REGION Network 6: 2 -Op2- - Reparare palete Zona A
   #f[#_op2](sA := #_nop0,   // "sta"
             nrs := #_op2,
             sB := #_cen,
             iA := "DB2_WORK_BITS".Transport_Conveyor_SQs.SQ_Repaired_Pallet[0] AND #tmr[5].Q,
             cEvac := NOT "x".evac[2],
             iAr := NOT "DB2_WORK_BITS".Transport_Conveyor_SQs.SQ_Repaired_Pallet[0],
             iB := "SCentrorMemT",
             cmdB => #tranzit[#_op2],
             ENO => #_w1);
   #f[2].condRetract := #_w1;
   #f[2].WrkDn := #_w1;
   #f[2].disAlm_apar := #_w1;
   #tmr[5].TON(IN := "DB2_WORK_BITS".Transport_Conveyor_SQs.SQ_Repaired_Pallet[0], PT := T#2s);
END_REGION

REGION Network 7: stoper op
   RUNG wire#powerrail
      Contact( "DB2_WORK_BITS".Transport_Conveyor_SQs.SQ_Repaired_Pallet[0] )
      wire#w1
      Coil( "O".StopReqUp1 )
   END_RUNG
   RUNG wire#powerrail
      Contact( #tranzit[#_op2] )
   END_RUNG wire#w1
   // the same network as SCL:
   "O".StopReqUp1 := "DB2_WORK_BITS".Transport_Conveyor_SQs.SQ_Repaired_Pallet[0] OR #tranzit[#_op2];
END_REGION

REGION Network 8
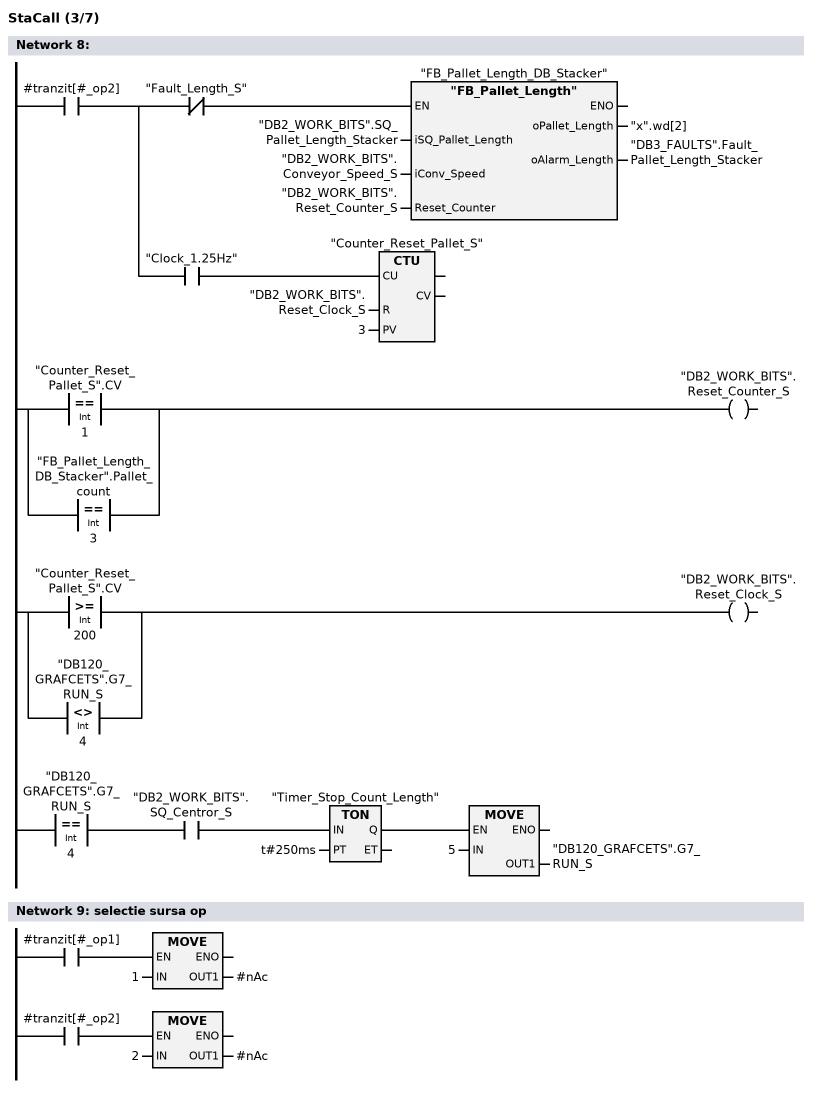
   IF #tranzit[#_op2] AND NOT "Fault_Length_S" THEN
       "FB_Pallet_Length_DB_Stacker"(iSQ_Pallet_Length := "DB2_WORK_BITS".SQ_Pallet_Length_Stacker,   // "FB_Pallet_Length"
                               iConv_Speed := "DB2_WORK_BITS".Conveyor_Speed_S,
                               Reset_Counter := "DB2_WORK_BITS".Reset_Counter_S,
                               oPallet_Length => "x".wd[2],
                               oAlarm_Length => "DB3_FAULTS".Fault_Pallet_Length_Stacker);
   END_IF;
   "Counter_Reset_Pallet_S".CTU(CU := #tranzit[#_op2] AND "Clock_1.25Hz",
                           R := "DB2_WORK_BITS".Reset_Clock_S,
                           PV := 3);
   "DB2_WORK_BITS".Reset_Counter_S := ("Counter_Reset_Pallet_S".CV = 1) OR ("FB_Pallet_Length_DB_Stacker".Pallet_count = 3);
   "DB2_WORK_BITS".Reset_Clock_S := ("Counter_Reset_Pallet_S".CV >= 200) OR ("DB120_GRAFCETS".G7_RUN_S <> 4);
   "Timer_Stop_Count_Length".TON(IN := ("DB120_GRAFCETS".G7_RUN_S = 4) AND "DB2_WORK_BITS".SQ_Centror_S,
                           PT := t#250ms);
   IF "Timer_Stop_Count_Length".Q THEN "DB120_GRAFCETS".G7_RUN_S := 5; END_IF;
END_REGION

REGION Network 9: selectie sursa op
   RUNG wire#powerrail
      Contact( #tranzit[#_op1] )
      Move(in := 1, out1 => #nAc)
   END_RUNG
   RUNG wire#powerrail
      Contact( #tranzit[#_op2] )
      Move(in := 2, out1 => #nAc)
   END_RUNG
   // the same network as SCL:
   IF #tranzit[#_op1] THEN #nAc := 1; END_IF;
   IF #tranzit[#_op2] THEN #nAc := 2; END_IF;
END_REGION

REGION Network 10: senz stop stk
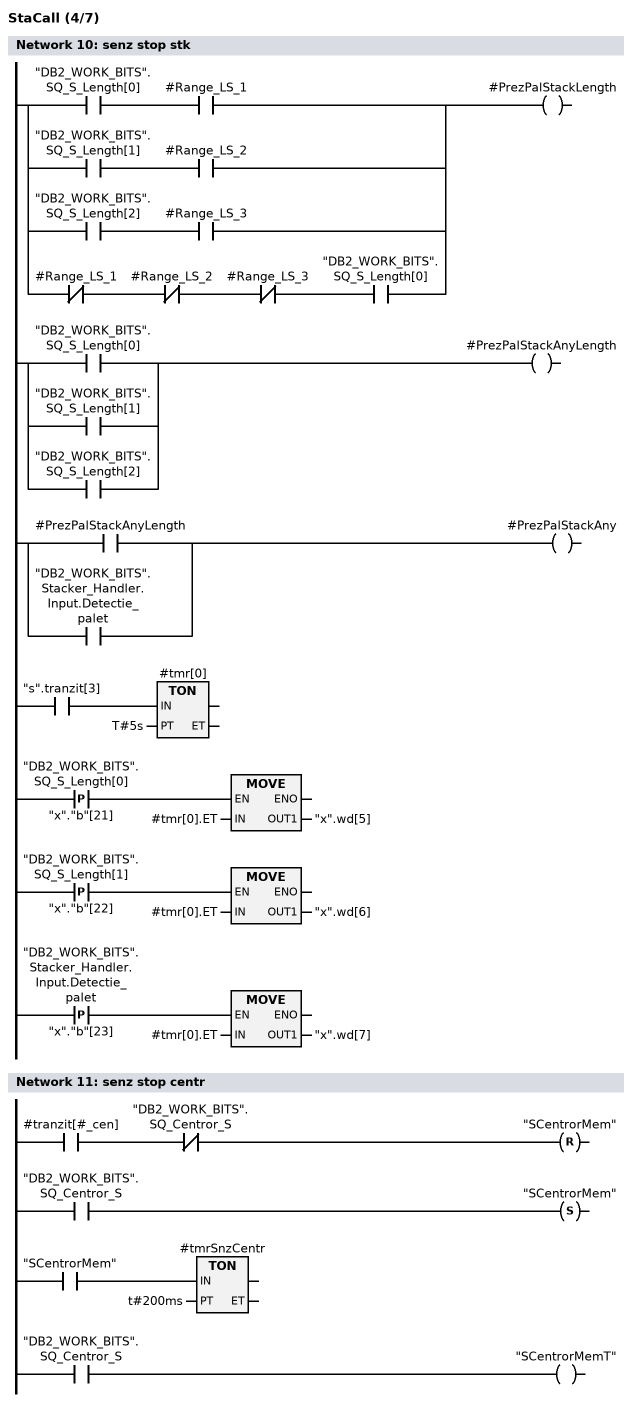
   #PrezPalStackLength := ("DB2_WORK_BITS".SQ_S_Length[0] AND #Range_LS_1) OR ("DB2_WORK_BITS".SQ_S_Length[1] AND #Range_LS_2) OR ("DB2_WORK_BITS".SQ_S_Length[2] AND #Range_LS_3) OR (NOT #Range_LS_1 AND NOT #Range_LS_2 AND NOT #Range_LS_3 AND "DB2_WORK_BITS".SQ_S_Length[0]);
   #PrezPalStackAnyLength := "DB2_WORK_BITS".SQ_S_Length[0] OR "DB2_WORK_BITS".SQ_S_Length[1] OR "DB2_WORK_BITS".SQ_S_Length[2];
   #PrezPalStackAny := #PrezPalStackAnyLength OR "DB2_WORK_BITS".Stacker_Handler.Input.Detectie_palet;
   #tmr[0].TON(IN := "s".tranzit[3], PT := T#5s);
   #_w1 := "DB2_WORK_BITS".SQ_S_Length[0] AND NOT "x"."b"[21];   // rising edge of "DB2_WORK_BITS".SQ_S_Length[0]
   "x"."b"[21] := "DB2_WORK_BITS".SQ_S_Length[0];
   IF #_w1 THEN "x".wd[5] := #tmr[0].ET; END_IF;
   #_w2 := "DB2_WORK_BITS".SQ_S_Length[1] AND NOT "x"."b"[22];   // rising edge of "DB2_WORK_BITS".SQ_S_Length[1]
   "x"."b"[22] := "DB2_WORK_BITS".SQ_S_Length[1];
   IF #_w2 THEN "x".wd[6] := #tmr[0].ET; END_IF;
   #_w3 := "DB2_WORK_BITS".Stacker_Handler.Input.Detectie_palet AND NOT "x"."b"[23];   // rising edge of "DB2_WORK_BITS".Stacker_Handler.Input.Detectie_palet
   "x"."b"[23] := "DB2_WORK_BITS".Stacker_Handler.Input.Detectie_palet;
   IF #_w3 THEN "x".wd[7] := #tmr[0].ET; END_IF;
END_REGION

REGION Network 11: senz stop centr
   IF #tranzit[#_cen] AND NOT "DB2_WORK_BITS".SQ_Centror_S THEN "SCentrorMem" := FALSE; END_IF;
   IF "DB2_WORK_BITS".SQ_Centror_S THEN "SCentrorMem" := TRUE; END_IF;
   #tmrSnzCentr(IN := "SCentrorMem", PT := t#200ms);   // TON
   "SCentrorMemT" := "DB2_WORK_BITS".SQ_Centror_S;
END_REGION

REGION Network 12: 3- Centror
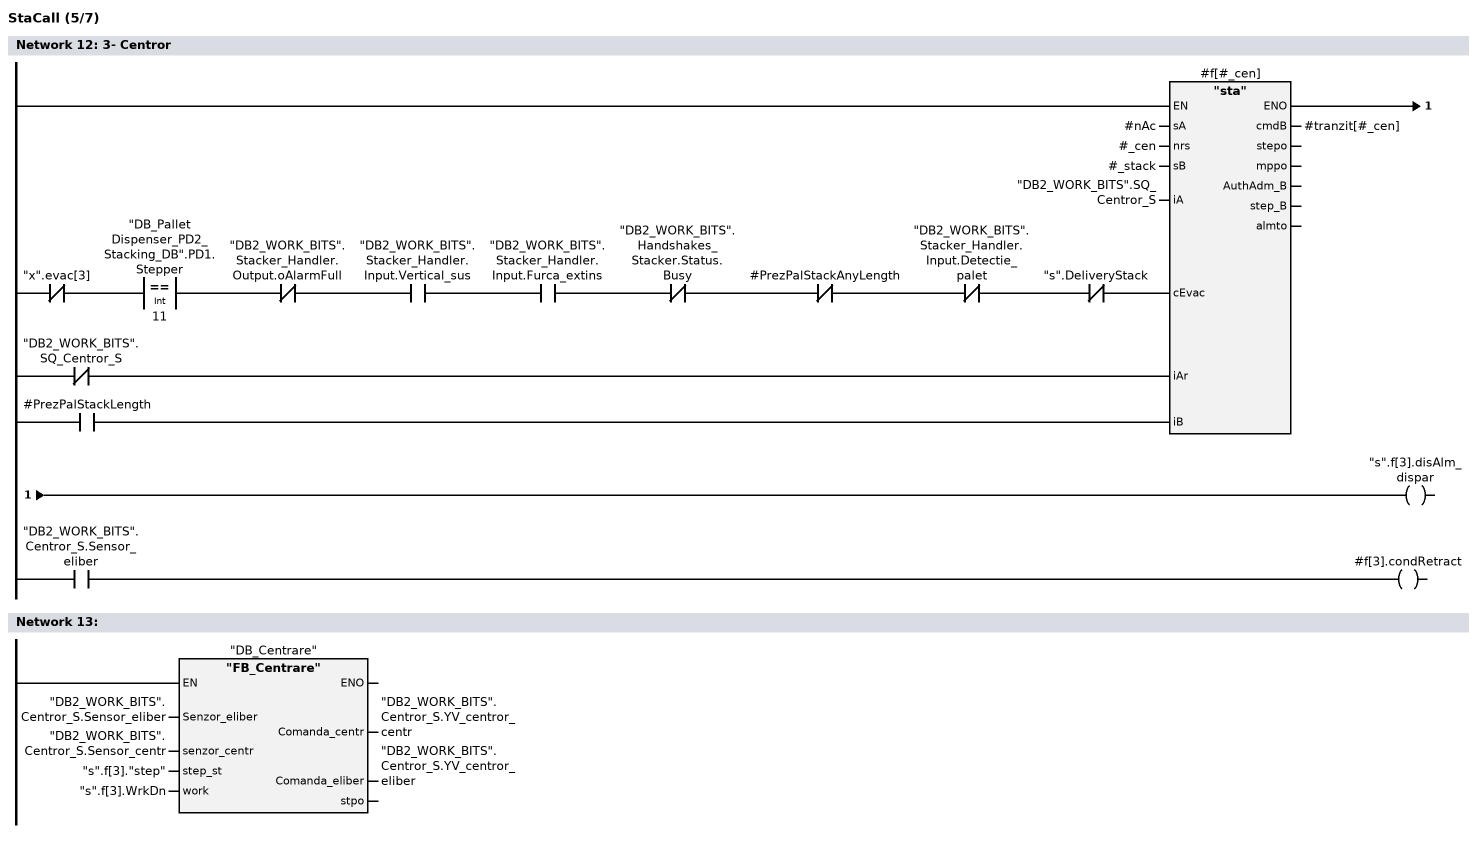
   RUNG wire#powerrail
      #f[#_cen](cEvac := wire#w1, iAr := wire#w2, iB := wire#w3, sA := #nAc, nrs := #_cen, sB := #_stack, iA := "DB2_WORK_BITS".SQ_Centror_S, cmdB => #tranzit[#_cen], stepo =>, mppo =>, AuthAdm_B =>, step_B =>, almto =>)
      Coil( "s".f[3].disAlm_dispar )
   END_RUNG
   RUNG wire#powerrail
      I_Contact( "x".evac[3] )
      { S7_Templates := "SrcType := Int" } EQ_Contact(in1 := "DB_PalletDispenser_PD2_Stacking_DB".PD1.Stepper, in2 := 11)
      I_Contact( "DB2_WORK_BITS".Stacker_Handler.Output.oAlarmFull )
      Contact( "DB2_WORK_BITS".Stacker_Handler.Input.Vertical_sus )
      Contact( "DB2_WORK_BITS".Stacker_Handler.Input.Furca_extins )
      I_Contact( "DB2_WORK_BITS".Handshakes_Stacker.Status.Busy )
      I_Contact( #PrezPalStackAnyLength )
      I_Contact( "DB2_WORK_BITS".Stacker_Handler.Input.Detectie_palet )
      I_Contact( "s".DeliveryStack )
   END_RUNG wire#w1
   RUNG wire#powerrail
      I_Contact( "DB2_WORK_BITS".SQ_Centror_S )
   END_RUNG wire#w2
   RUNG wire#powerrail
      Contact( #PrezPalStackLength )
   END_RUNG wire#w3
   RUNG wire#powerrail
      Contact( "DB2_WORK_BITS".Centror_S.Sensor_eliber )
      Coil( #f[3].condRetract )
   END_RUNG
   // the same network as SCL:
   #f[#_cen](sA := #nAc,   // "sta"
             nrs := #_cen,
             sB := #_stack,
             iA := "DB2_WORK_BITS".SQ_Centror_S,
             cEvac := NOT "x".evac[3] AND ("DB_PalletDispenser_PD2_Stacking_DB".PD1.Stepper = 11) AND NOT "DB2_WORK_BITS".Stacker_Handler.Output.oAlarmFull AND "DB2_WORK_BITS".Stacker_Handler.Input.Vertical_sus AND "DB2_WORK_BITS".Stacker_Handler.Input.Furca_extins AND NOT "DB2_WORK_BITS".Handshakes_Stacker.Status.Busy AND NOT #PrezPalStackAnyLength AND NOT "DB2_WORK_BITS".Stacker_Handler.Input.Detectie_palet AND NOT "s".DeliveryStack,
             iAr := NOT "DB2_WORK_BITS".SQ_Centror_S,
             iB := #PrezPalStackLength,
             cmdB => #tranzit[#_cen],
             ENO => #_w1);
   "s".f[3].disAlm_dispar := #_w1;
   #f[3].condRetract := "DB2_WORK_BITS".Centror_S.Sensor_eliber;
END_REGION

REGION Network 13
   RUNG wire#powerrail
      "DB_Centrare"(Senzor_eliber := "DB2_WORK_BITS".Centror_S.Sensor_eliber, senzor_centr := "DB2_WORK_BITS".Centror_S.Sensor_centr, step_st := "s".f[3]."step", work := "s".f[3].WrkDn, Comanda_centr => "DB2_WORK_BITS".Centror_S.YV_centror_centr, Comanda_eliber => "DB2_WORK_BITS".Centror_S.YV_centror_eliber, stpo =>)
   END_RUNG
   // the same network as SCL:
   "DB_Centrare"(Senzor_eliber := "DB2_WORK_BITS".Centror_S.Sensor_eliber,   // "FB_Centrare"
                 senzor_centr := "DB2_WORK_BITS".Centror_S.Sensor_centr,
                 step_st := "s".f[3]."step",
                 work := "s".f[3].WrkDn,
                 Comanda_centr => "DB2_WORK_BITS".Centror_S.YV_centror_centr,
                 Comanda_eliber => "DB2_WORK_BITS".Centror_S.YV_centror_eliber);
END_REGION

REGION Network 14: 4- stacker
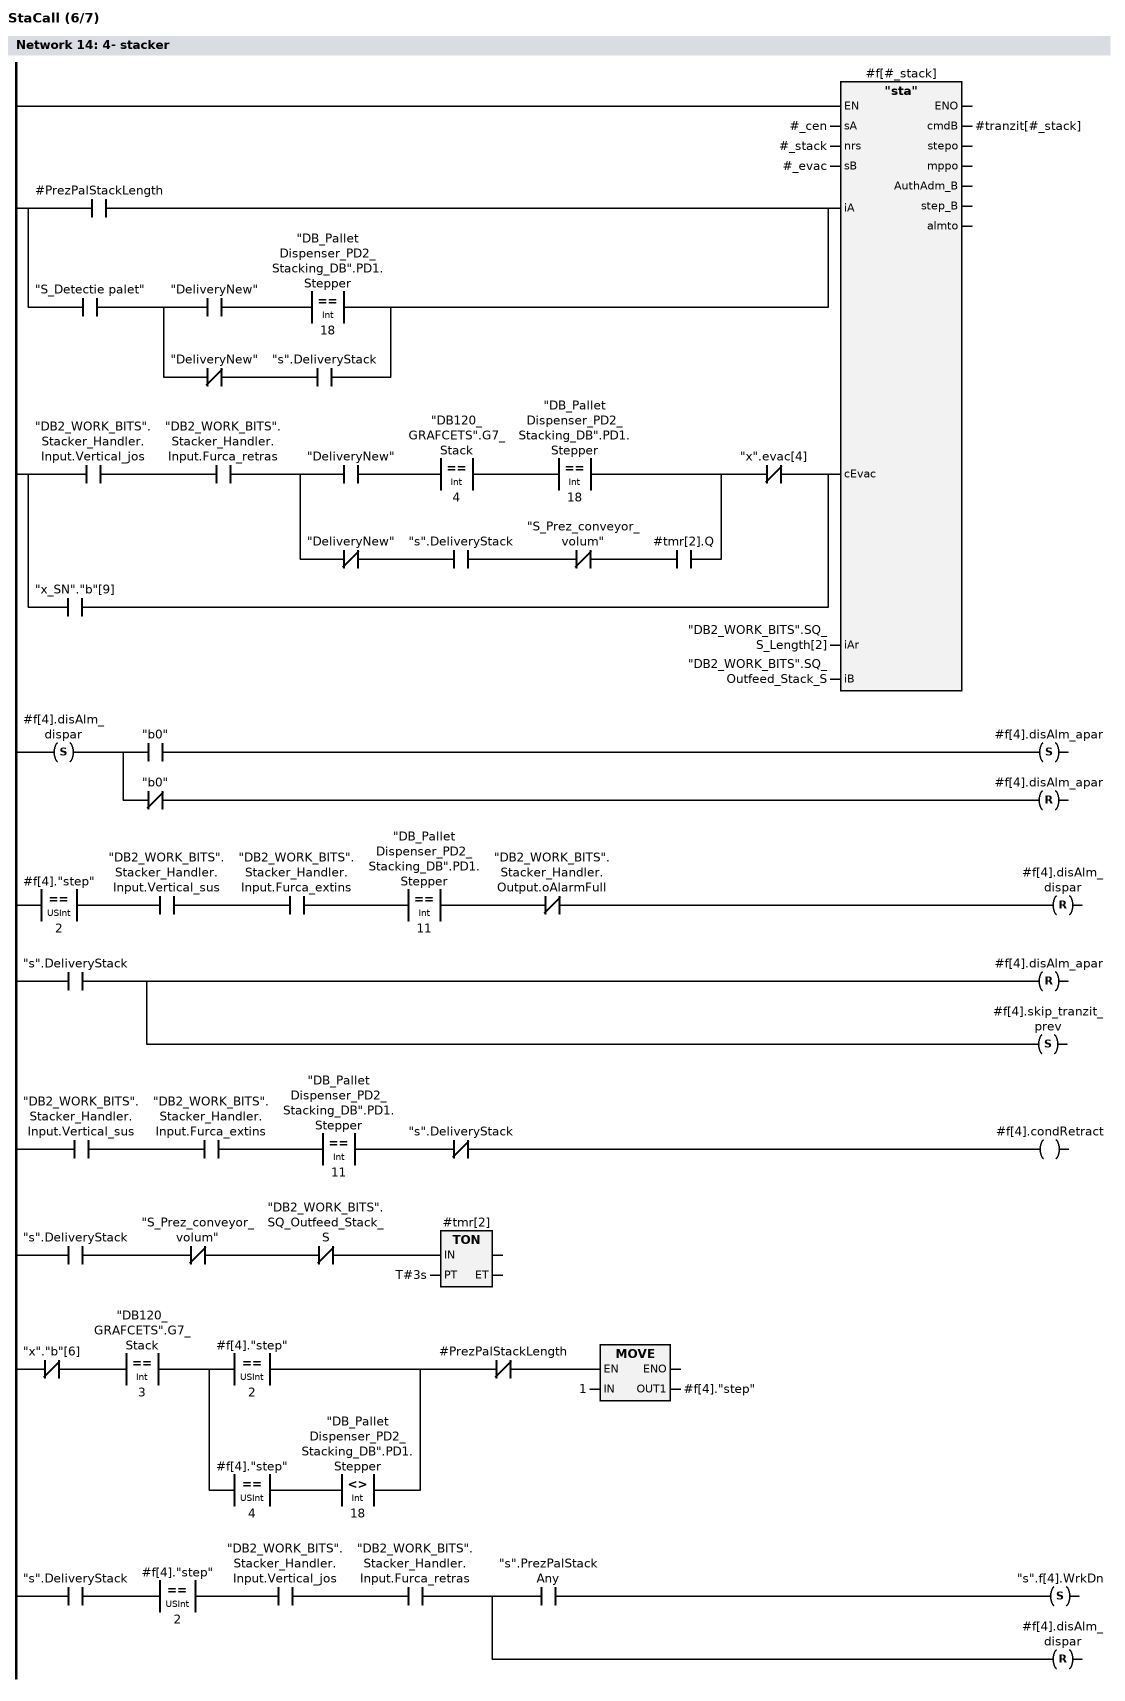
   #f[#_stack](sA := #_cen,   // "sta"
               nrs := #_stack,
               sB := #_evac,
               iA := #PrezPalStackLength OR ("S_Detectie palet" AND (("DeliveryNew" AND ("DB_PalletDispenser_PD2_Stacking_DB".PD1.Stepper = 18)) OR (NOT "DeliveryNew" AND "s".DeliveryStack))),
               cEvac := ("DB2_WORK_BITS".Stacker_Handler.Input.Vertical_jos AND "DB2_WORK_BITS".Stacker_Handler.Input.Furca_retras AND (("DeliveryNew" AND ("DB120_GRAFCETS".G7_Stack = 4) AND ("DB_PalletDispenser_PD2_Stacking_DB".PD1.Stepper = 18)) OR (NOT "DeliveryNew" AND "s".DeliveryStack AND NOT "S_Prez_conveyor_volum" AND #tmr[2].Q)) AND NOT "x".evac[4]) OR "x_SN"."b"[9],
               iAr := "DB2_WORK_BITS".SQ_S_Length[2],
               iB := "DB2_WORK_BITS".SQ_Outfeed_Stack_S,
               cmdB => #tranzit[#_stack]);
   #f[4].disAlm_dispar := TRUE;
   IF "b0" THEN #f[4].disAlm_apar := TRUE; END_IF;
   IF NOT "b0" THEN #f[4].disAlm_apar := FALSE; END_IF;
   IF (#f[4]."step" = 2) AND "DB2_WORK_BITS".Stacker_Handler.Input.Vertical_sus AND "DB2_WORK_BITS".Stacker_Handler.Input.Furca_extins AND ("DB_PalletDispenser_PD2_Stacking_DB".PD1.Stepper = 11) AND NOT "DB2_WORK_BITS".Stacker_Handler.Output.oAlarmFull THEN
       #f[4].disAlm_dispar := FALSE;
   END_IF;
   IF "s".DeliveryStack THEN
       #f[4].disAlm_apar := FALSE;
       #f[4].skip_tranzit_prev := TRUE;
   END_IF;
   #f[4].condRetract := "DB2_WORK_BITS".Stacker_Handler.Input.Vertical_sus AND "DB2_WORK_BITS".Stacker_Handler.Input.Furca_extins AND ("DB_PalletDispenser_PD2_Stacking_DB".PD1.Stepper = 11) AND NOT "s".DeliveryStack;
   #tmr[2].TON(IN := "s".DeliveryStack AND NOT "S_Prez_conveyor_volum" AND NOT "DB2_WORK_BITS".SQ_Outfeed_Stack_S,
               PT := T#3s);
   IF NOT "x"."b"[6] AND ("DB120_GRAFCETS".G7_Stack = 3) AND ((#f[4]."step" = 2) OR ((#f[4]."step" = 4) AND ("DB_PalletDispenser_PD2_Stacking_DB".PD1.Stepper <> 18))) AND NOT #PrezPalStackLength THEN
       #f[4]."step" := 1;
   END_IF;
   #_w1 := "s".DeliveryStack AND (#f[4]."step" = 2) AND "DB2_WORK_BITS".Stacker_Handler.Input.Vertical_jos AND "DB2_WORK_BITS".Stacker_Handler.Input.Furca_retras;
   IF #_w1 AND "s".PrezPalStackAny THEN "s".f[4].WrkDn := TRUE; END_IF;
   IF #_w1 THEN #f[4].disAlm_dispar := FALSE; END_IF;
END_REGION

REGION Network 15: 5- evac
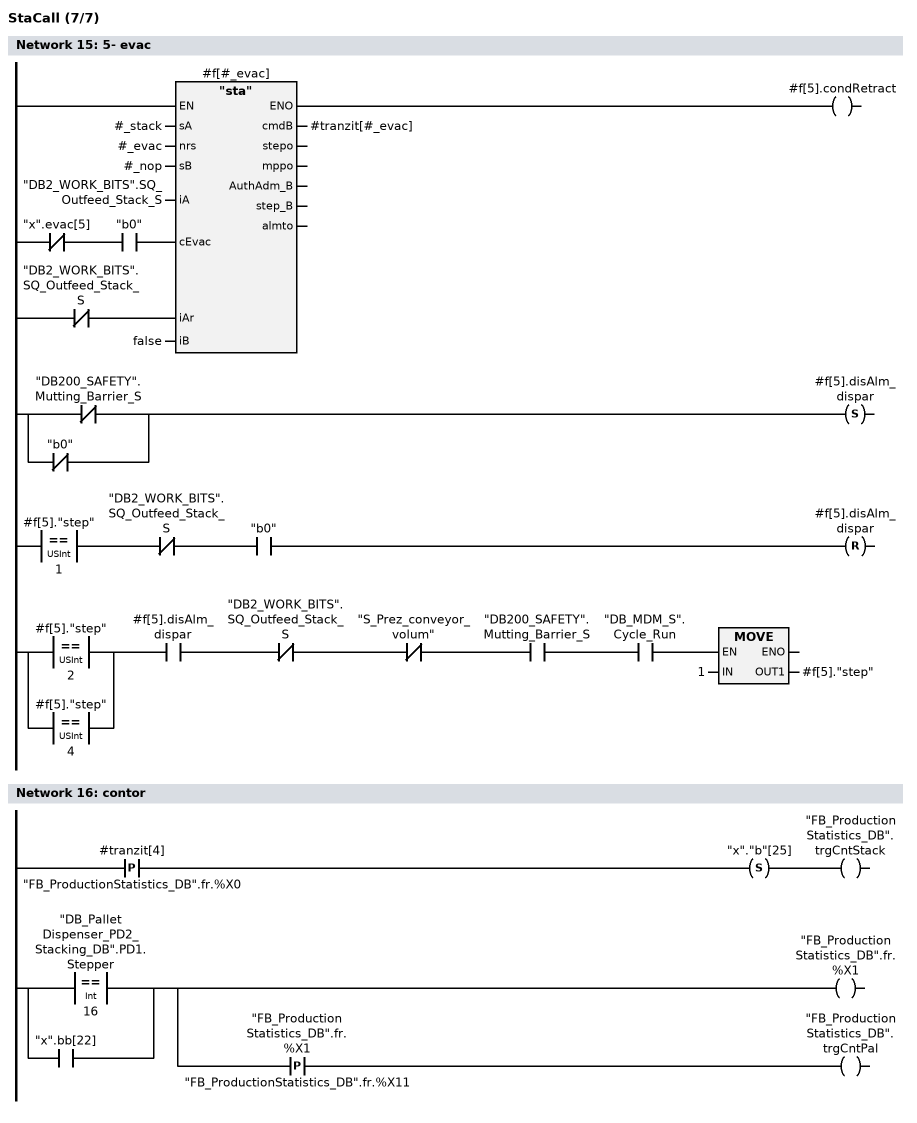
   RUNG wire#powerrail
      #f[#_evac](cEvac := wire#w1, iAr := wire#w2, sA := #_stack, nrs := #_evac, sB := #_nop, iA := "DB2_WORK_BITS".SQ_Outfeed_Stack_S, iB := false, cmdB => #tranzit[#_evac], stepo =>, mppo =>, AuthAdm_B =>, step_B =>, almto =>)
      Coil( #f[5].condRetract )
   END_RUNG
   RUNG wire#powerrail
      I_Contact( "x".evac[5] )
      Contact( "b0" )
   END_RUNG wire#w1
   RUNG wire#powerrail
      I_Contact( "DB2_WORK_BITS".SQ_Outfeed_Stack_S )
   END_RUNG wire#w2
   RUNG wire#powerrail
      I_Contact( "DB200_SAFETY".Mutting_Barrier_S )
      wire#w3
      S_Coil( #f[5].disAlm_dispar )
   END_RUNG
   RUNG wire#powerrail
      I_Contact( "b0" )
   END_RUNG wire#w3
   RUNG wire#powerrail
      { S7_Templates := "SrcType := USInt" } EQ_Contact(in1 := #f[5]."step", in2 := 1)
      I_Contact( "DB2_WORK_BITS".SQ_Outfeed_Stack_S )
      Contact( "b0" )
      R_Coil( #f[5].disAlm_dispar )
   END_RUNG
   RUNG wire#powerrail
      { S7_Templates := "SrcType := USInt" } EQ_Contact(in1 := #f[5]."step", in2 := 2)
      wire#w4
      Contact( #f[5].disAlm_dispar )
      I_Contact( "DB2_WORK_BITS".SQ_Outfeed_Stack_S )
      I_Contact( "S_Prez_conveyor_volum" )
      Contact( "DB200_SAFETY".Mutting_Barrier_S )
      Contact( "DB_MDM_S".Cycle_Run )
      Move(in := 1, out1 => #f[5]."step")
   END_RUNG
   RUNG wire#powerrail
      { S7_Templates := "SrcType := USInt" } EQ_Contact(in1 := #f[5]."step", in2 := 4)
   END_RUNG wire#w4
   // the same network as SCL:
   #f[#_evac](sA := #_stack,   // "sta"
              nrs := #_evac,
              sB := #_nop,
              iA := "DB2_WORK_BITS".SQ_Outfeed_Stack_S,
              cEvac := NOT "x".evac[5] AND "b0",
              iAr := NOT "DB2_WORK_BITS".SQ_Outfeed_Stack_S,
              iB := false,
              cmdB => #tranzit[#_evac],
              ENO => #_w1);
   #f[5].condRetract := #_w1;
   IF NOT "DB200_SAFETY".Mutting_Barrier_S OR NOT "b0" THEN #f[5].disAlm_dispar := TRUE; END_IF;
   IF (#f[5]."step" = 1) AND NOT "DB2_WORK_BITS".SQ_Outfeed_Stack_S AND "b0" THEN
       #f[5].disAlm_dispar := FALSE;
   END_IF;
   IF ((#f[5]."step" = 2) OR (#f[5]."step" = 4)) AND #f[5].disAlm_dispar AND NOT "DB2_WORK_BITS".SQ_Outfeed_Stack_S AND NOT "S_Prez_conveyor_volum" AND "DB200_SAFETY".Mutting_Barrier_S AND "DB_MDM_S".Cycle_Run THEN
       #f[5]."step" := 1;
   END_IF;
END_REGION

REGION Network 16: contor
   RUNG wire#powerrail
      P_Contact(operand := #tranzit[4], bit := "FB_ProductionStatistics_DB".fr.%X0)
      S_Coil( "x"."b"[25] )
      Coil( "FB_ProductionStatistics_DB".trgCntStack )
   END_RUNG
   RUNG wire#powerrail
      { S7_Templates := "SrcType := Int" } EQ_Contact(in1 := "DB_PalletDispenser_PD2_Stacking_DB".PD1.Stepper, in2 := 16)
      wire#w1
      Coil( "FB_ProductionStatistics_DB".fr.%X1 )
   END_RUNG
   RUNG wire#powerrail
      Contact( "x".bb[22] )
   END_RUNG wire#w1
   RUNG wire#w1
      P_Contact(operand := "FB_ProductionStatistics_DB".fr.%X1, bit := "FB_ProductionStatistics_DB".fr.%X11)
      Coil( "FB_ProductionStatistics_DB".trgCntPal )
   END_RUNG
   // the same network as SCL:
   #_w1 := #tranzit[4] AND NOT "FB_ProductionStatistics_DB".fr.%X0;   // rising edge of #tranzit[4]
   "FB_ProductionStatistics_DB".fr.%X0 := #tranzit[4];
   IF #_w1 THEN "x"."b"[25] := TRUE; END_IF;
   "FB_ProductionStatistics_DB".trgCntStack := #_w1;
   "FB_ProductionStatistics_DB".fr.%X1 := ("DB_PalletDispenser_PD2_Stacking_DB".PD1.Stepper = 16) OR "x".bb[22];
   #_w2 := "FB_ProductionStatistics_DB".fr.%X1 AND "FB_ProductionStatistics_DB".fr.%X1 AND NOT "FB_ProductionStatistics_DB".fr.%X11;   // rising edge of "FB_ProductionStatistics_DB".fr.%X1
   "FB_ProductionStatistics_DB".fr.%X11 := "FB_ProductionStatistics_DB".fr.%X1;
   "FB_ProductionStatistics_DB".trgCntPal := #_w2;
END_REGION
END_FUNCTION_BLOCK

FUNCTION_BLOCK "sta"   // FB13, LAD
{ S7_Optimized_Access := 'TRUE' }
VERSION : 0.1
   VAR_INPUT
      sA : USInt;   // statie Admit
      nrs : USInt;   // statie crt
      sB : USInt;   // statie Evac
      iA : Bool;   // conditie Admit
      cEvac : Bool;
      iAr : Bool;   // cond Release
      iB : Bool;   // cond Evac
   END_VAR
   VAR_OUTPUT
      cmdB : Bool;
      stepo : USInt;
      mppo : Bool;
      AuthAdm_B : Bool;
      step_B : USInt;
      almto : USInt;
   END_VAR
   VAR
      "step" : USInt;
      stepv : USInt;
      mpp : Bool;
      alm_apar : Bool;
      alm_disapear : Bool;
      alm_tmt : Bool;
      alm_release : Bool;
      AuthAdmit : Bool;
      AuthEvacEx : Bool;
      almt : Bool;
      WrkDn : Bool;
      condRetract : Bool;
      skip_tranzit_prev : Bool;
      product_disapear_confirmed : Bool;
      transit_end_confirmed : Bool;
      tim_alm : Array[1..6] of IEC_TIMER;
      HMI_stat_s : USInt;
      disAlm_Tmt : Bool;
      disAlm_dispar : Bool;
      disAlm_apar : Bool;
      disAlmRls : Bool;
      HMI_stat_t : USInt;
      tranzit_mem : Bool;
      cycle : Bool;
      almw : Word;
      HMI_statT : USInt;
      HMI_statS : USInt;
      tr : USInt;
      AlarmW : Word;
   END_VAR
   VAR_TEMP
      tmpui : SInt;
   END_VAR
   VAR CONSTANT
      b0 : Bool;
   END_VAR
   VAR_TEMP   // added for the SCL form of the ladder/FBD networks
      _w1 : Bool;
      _w2 : Bool;
      _w3 : Bool;
   END_VAR
BEGIN

REGION Network 1: first cycle
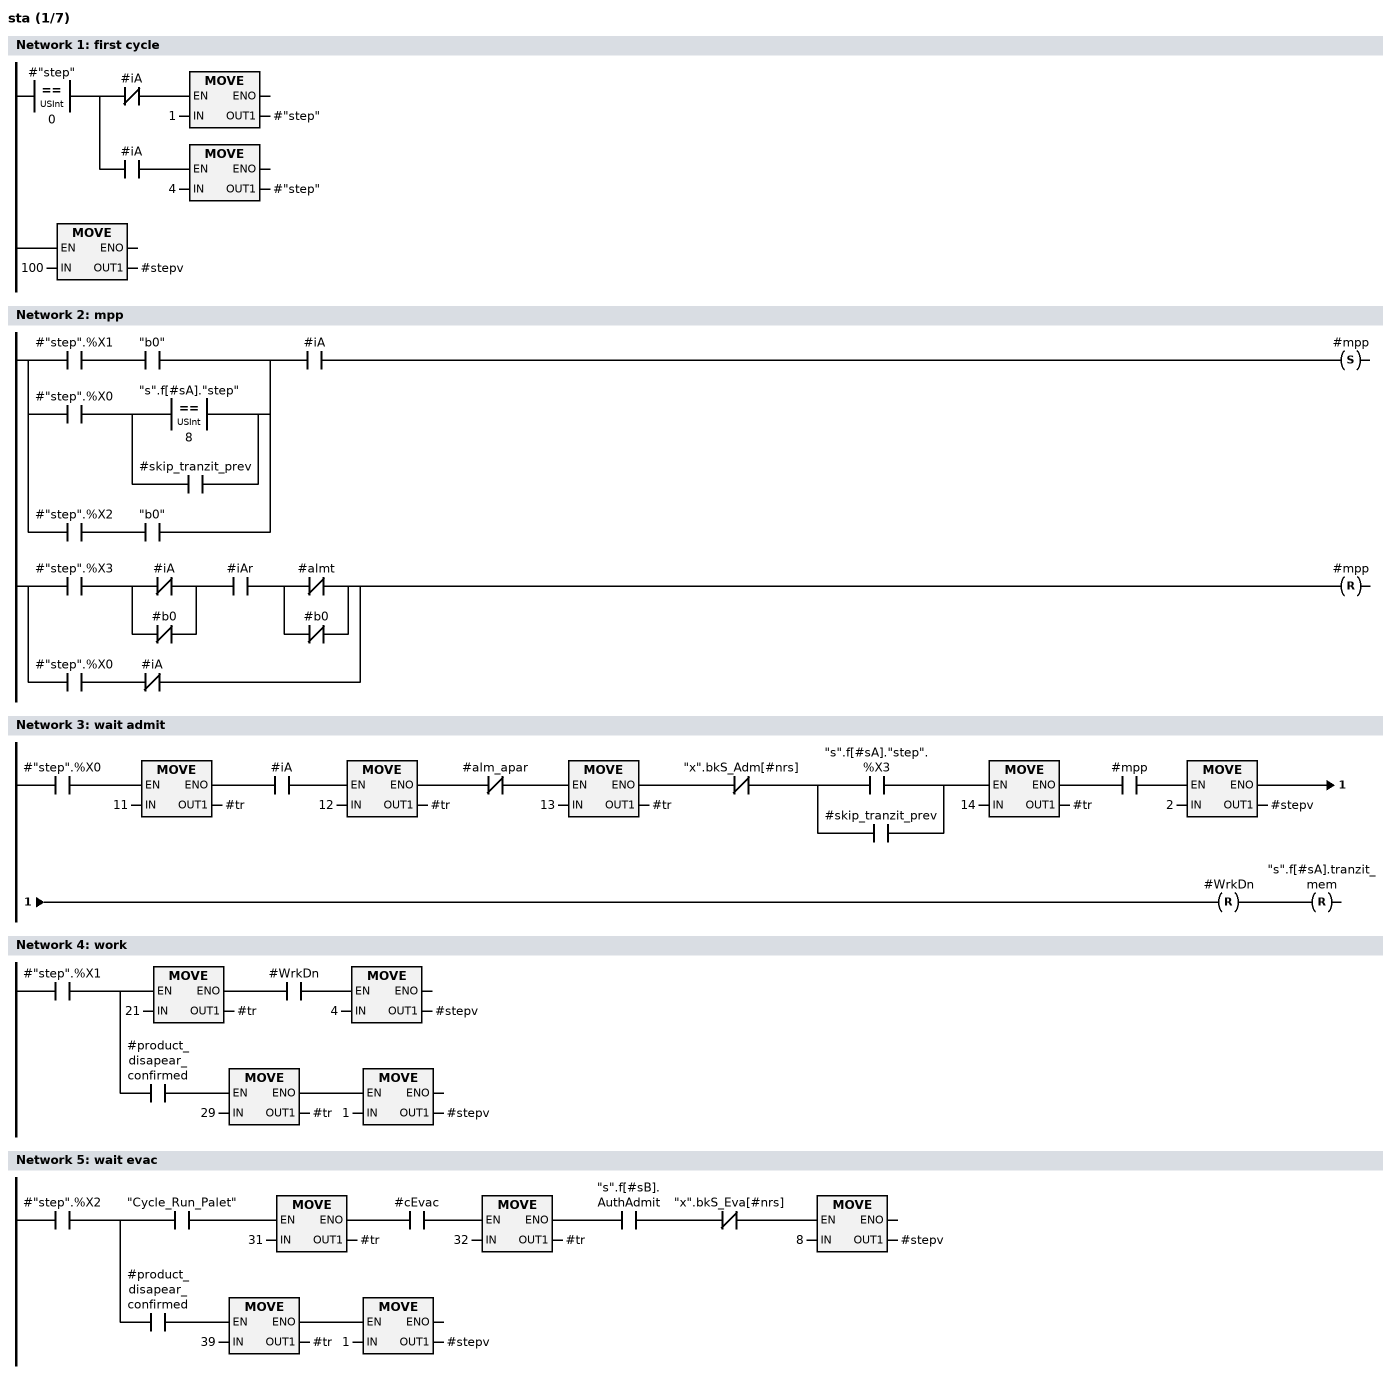
   RUNG wire#powerrail
      { S7_Templates := "SrcType := USInt" } EQ_Contact(in1 := #"step", in2 := 0)
      wire#w1
      I_Contact( #iA )
      Move(in := 1, out1 => #"step")
   END_RUNG
   RUNG wire#w1
      Contact( #iA )
      Move(in := 4, out1 => #"step")
   END_RUNG
   RUNG wire#powerrail
      Move(in := 100, out1 => #stepv)
   END_RUNG
   // the same network as SCL:
   #_w1 := #"step" = 0;
   IF #_w1 AND NOT #iA THEN #"step" := 1; END_IF;
   IF #_w1 AND #iA THEN #"step" := 4; END_IF;
   #stepv := 100;
END_REGION

REGION Network 2: mpp
   RUNG wire#powerrail
      Contact( #"step".%X1 )
      Contact( "b0" )
      wire#w1
      Contact( #iA )
      S_Coil( #mpp )
   END_RUNG
   RUNG wire#powerrail
      Contact( #"step".%X0 )
      wire#w2
      { S7_Templates := "SrcType := USInt" } EQ_Contact(in1 := "s".f[#sA]."step", in2 := 8)
   END_RUNG wire#w1
   RUNG wire#w2
      Contact( #skip_tranzit_prev )
   END_RUNG wire#w1
   RUNG wire#powerrail
      Contact( #"step".%X2 )
      Contact( "b0" )
   END_RUNG wire#w1
   RUNG wire#powerrail
      Contact( #"step".%X3 )
      wire#w3
      I_Contact( #iA )
      wire#w4
      Contact( #iAr )
      wire#w5
      I_Contact( #almt )
      wire#w6
      R_Coil( #mpp )
   END_RUNG
   RUNG wire#w3
      I_Contact( #b0 )
   END_RUNG wire#w4
   RUNG wire#w5
      I_Contact( #b0 )
   END_RUNG wire#w6
   RUNG wire#powerrail
      Contact( #"step".%X0 )
      I_Contact( #iA )
   END_RUNG wire#w6
   // the same network as SCL:
   IF ((#"step".%X1 AND "b0") OR (#"step".%X0 AND (("s".f[#sA]."step" = 8) OR #skip_tranzit_prev)) OR (#"step".%X2 AND "b0")) AND #iA THEN
       #mpp := TRUE;
   END_IF;
   IF (#"step".%X3 AND (NOT #iA OR NOT #b0) AND #iAr AND (NOT #almt OR NOT #b0)) OR (#"step".%X0 AND NOT #iA) THEN
       #mpp := FALSE;
   END_IF;
END_REGION

REGION Network 3: wait admit
   RUNG wire#powerrail
      Contact( #"step".%X0 )
      Move(in := 11, out1 => #tr)
      Contact( #iA )
      Move(in := 12, out1 => #tr)
      I_Contact( #alm_apar )
      Move(in := 13, out1 => #tr)
      I_Contact( "x".bkS_Adm[#nrs] )
      wire#w1
      Contact( "s".f[#sA]."step".%X3 )
      wire#w2
      Move(in := 14, out1 => #tr)
      Contact( #mpp )
      Move(in := 2, out1 => #stepv)
      R_Coil( #WrkDn )
      R_Coil( "s".f[#sA].tranzit_mem )
   END_RUNG
   RUNG wire#w1
      Contact( #skip_tranzit_prev )
   END_RUNG wire#w2
   // the same network as SCL:
   IF #"step".%X0 THEN #tr := 11; END_IF;
   #_w1 := #"step".%X0 AND #iA;
   IF #_w1 THEN #tr := 12; END_IF;
   #_w2 := #_w1 AND NOT #alm_apar;
   IF #_w2 THEN #tr := 13; END_IF;
   #_w3 := #_w2 AND NOT "x".bkS_Adm[#nrs] AND ("s".f[#sA]."step".%X3 OR #skip_tranzit_prev);
   IF #_w3 THEN #tr := 14; END_IF;
   IF #_w3 AND #mpp THEN
       #stepv := 2;
       #WrkDn := FALSE;
       "s".f[#sA].tranzit_mem := FALSE;
   END_IF;
END_REGION

REGION Network 4: work
   RUNG wire#powerrail
      Contact( #"step".%X1 )
      wire#w1
      Move(in := 21, out1 => #tr)
      Contact( #WrkDn )
      Move(in := 4, out1 => #stepv)
   END_RUNG
   RUNG wire#w1
      Contact( #product_disapear_confirmed )
      Move(in := 29, out1 => #tr)
      Move(in := 1, out1 => #stepv)
   END_RUNG
   // the same network as SCL:
   IF #"step".%X1 THEN #tr := 21; END_IF;
   IF #"step".%X1 AND #WrkDn THEN #stepv := 4; END_IF;
   IF #"step".%X1 AND #product_disapear_confirmed THEN
       #tr := 29;
       #stepv := 1;
   END_IF;
END_REGION

REGION Network 5: wait evac
   RUNG wire#powerrail
      Contact( #"step".%X2 )
      wire#w1
      Contact( "Cycle_Run_Palet" )
      Move(in := 31, out1 => #tr)
      Contact( #cEvac )
      Move(in := 32, out1 => #tr)
      Contact( "s".f[#sB].AuthAdmit )
      I_Contact( "x".bkS_Eva[#nrs] )
      Move(in := 8, out1 => #stepv)
   END_RUNG
   RUNG wire#w1
      Contact( #product_disapear_confirmed )
      Move(in := 39, out1 => #tr)
      Move(in := 1, out1 => #stepv)
   END_RUNG
   // the same network as SCL:
   #_w1 := #"step".%X2 AND "Cycle_Run_Palet";
   IF #_w1 THEN #tr := 31; END_IF;
   #_w2 := #_w1 AND #cEvac;
   IF #_w2 THEN #tr := 32; END_IF;
   IF #_w2 AND "s".f[#sB].AuthAdmit AND NOT "x".bkS_Eva[#nrs] THEN #stepv := 8; END_IF;
   IF #"step".%X2 AND #product_disapear_confirmed THEN
       #tr := 39;
       #stepv := 1;
   END_IF;
END_REGION

REGION Network 6: evac